(* Logix 5000 project; controller _GigaDiscovery vendor 1 type 14 code 244 rev 35.11; software revision 35.03; part 17 of 23 *)
(* tags used below, declared in another part *)
   Os : DINT;
   All_Rack_Left_Sensor_FP_OFF : BOOL;
   All_Rack_Left_Sensor_O1_OFF : BOOL;
   All_Rack_Right_Sensor_FP_OFF : BOOL;
   All_Rack_Right_Sensor_O1_OFF : BOOL;
   All_Rack_Sensor_OFF : BOOL;
   Mem_All_Rack_Sensor_OFF : BOOL;
   OS_Start_Stop_Cycle_Started : BOOL;
   Reset_Pulse : BOOL;
   RESTRAINTS_Closed : BOOL;   // All RESTRAINTS Closed
   Restraints_Cycle : Sequencer;
   RESTRAINTS_Rack : LapBar_Racks[41];
   RESTRAINTS_Rack_Sector_ON : BOOL;
   RESTRAINTS_Sector : LapBars_Sector[9];
   Start_Autom_Cycle : Sequencer;
   Start_Stop_Cycle : Sequencer;
(* S_Input, continued *)

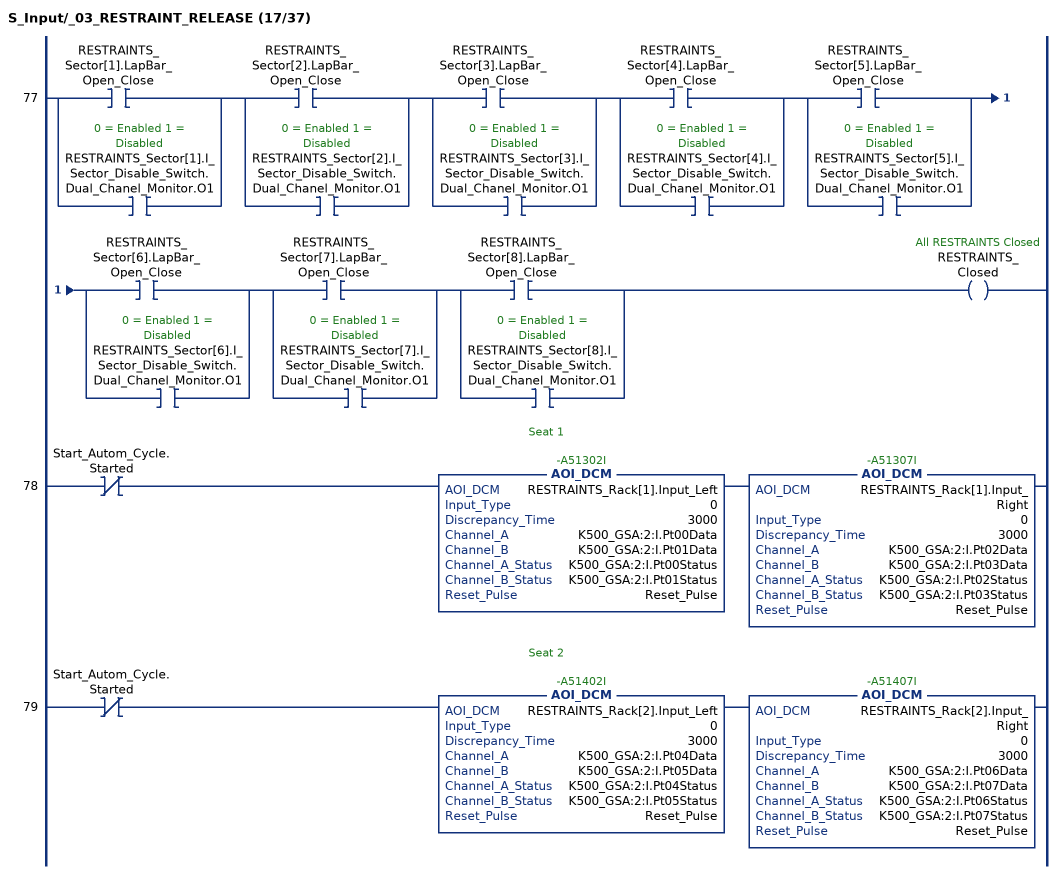
   [picture p324: S_Input/_03_RESTRAINT_RELEASE rungs 77-79]
   77: [XIC(RESTRAINTS_Sector[1].LapBar_Open_Close) ,XIC(RESTRAINTS_Sector[1].I_Sector_Disable_Switch.Dual_Chanel_Monitor.O1) ][XIC(RESTRAINTS_Sector[2].LapBar_Open_Close) ,XIC(RESTRAINTS_Sector[2].I_Sector_Disable_Switch.Dual_Chanel_Monitor.O1) ][XIC(RESTRAINTS_Sector[3].LapBar_Open_Close) ,XIC(RESTRAINTS_Sector[3].I_Sector_Disable_Switch.Dual_Chanel_Monitor.O1) ][XIC(RESTRAINTS_Sector[4].LapBar_Open_Close) ,XIC(RESTRAINTS_Sector[4].I_Sector_Disable_Switch.Dual_Chanel_Monitor.O1) ][XIC(RESTRAINTS_Sector[5].LapBar_Open_Close) ,XIC(RESTRAINTS_Sector[5].I_Sector_Disable_Switch.Dual_Chanel_Monitor.O1) ][XIC(RESTRAINTS_Sector[6].LapBar_Open_Close) ,XIC(RESTRAINTS_Sector[6].I_Sector_Disable_Switch.Dual_Chanel_Monitor.O1) ][XIC(RESTRAINTS_Sector[7].LapBar_Open_Close) ,XIC(RESTRAINTS_Sector[7].I_Sector_Disable_Switch.Dual_Chanel_Monitor.O1) ][XIC(RESTRAINTS_Sector[8].LapBar_Open_Close) ,XIC(RESTRAINTS_Sector[8].I_Sector_Disable_Switch.Dual_Chanel_Monitor.O1) ]OTE(RESTRAINTS_Closed);
   // Seat 1
   78: XIO(Start_Autom_Cycle.Started)AOI_DCM(RESTRAINTS_Rack[1].Input_Left,0,3000,K500_GSA:2:I.Pt00Data,K500_GSA:2:I.Pt01Data,K500_GSA:2:I.Pt00Status,K500_GSA:2:I.Pt01Status,Reset_Pulse)AOI_DCM(RESTRAINTS_Rack[1].Input_Right,0,3000,K500_GSA:2:I.Pt02Data,K500_GSA:2:I.Pt03Data,K500_GSA:2:I.Pt02Status,K500_GSA:2:I.Pt03Status,Reset_Pulse);
   // Seat 2
   79: XIO(Start_Autom_Cycle.Started)AOI_DCM(RESTRAINTS_Rack[2].Input_Left,0,3000,K500_GSA:2:I.Pt04Data,K500_GSA:2:I.Pt05Data,K500_GSA:2:I.Pt04Status,K500_GSA:2:I.Pt05Status,Reset_Pulse)AOI_DCM(RESTRAINTS_Rack[2].Input_Right,0,3000,K500_GSA:2:I.Pt06Data,K500_GSA:2:I.Pt07Data,K500_GSA:2:I.Pt06Status,K500_GSA:2:I.Pt07Status,Reset_Pulse);
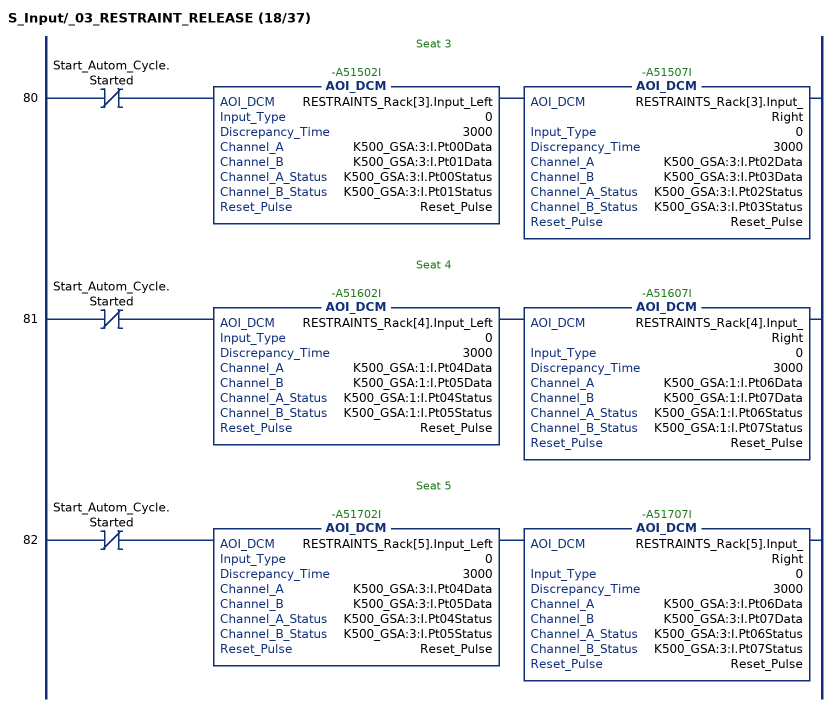
   // Seat 3
   80: XIO(Start_Autom_Cycle.Started)AOI_DCM(RESTRAINTS_Rack[3].Input_Left,0,3000,K500_GSA:3:I.Pt00Data,K500_GSA:3:I.Pt01Data,K500_GSA:3:I.Pt00Status,K500_GSA:3:I.Pt01Status,Reset_Pulse)AOI_DCM(RESTRAINTS_Rack[3].Input_Right,0,3000,K500_GSA:3:I.Pt02Data,K500_GSA:3:I.Pt03Data,K500_GSA:3:I.Pt02Status,K500_GSA:3:I.Pt03Status,Reset_Pulse);
   // Seat 4
   81: XIO(Start_Autom_Cycle.Started)AOI_DCM(RESTRAINTS_Rack[4].Input_Left,0,3000,K500_GSA:1:I.Pt04Data,K500_GSA:1:I.Pt05Data,K500_GSA:1:I.Pt04Status,K500_GSA:1:I.Pt05Status,Reset_Pulse)AOI_DCM(RESTRAINTS_Rack[4].Input_Right,0,3000,K500_GSA:1:I.Pt06Data,K500_GSA:1:I.Pt07Data,K500_GSA:1:I.Pt06Status,K500_GSA:1:I.Pt07Status,Reset_Pulse);
   // Seat 5
   82: XIO(Start_Autom_Cycle.Started)AOI_DCM(RESTRAINTS_Rack[5].Input_Left,0,3000,K500_GSA:3:I.Pt04Data,K500_GSA:3:I.Pt05Data,K500_GSA:3:I.Pt04Status,K500_GSA:3:I.Pt05Status,Reset_Pulse)AOI_DCM(RESTRAINTS_Rack[5].Input_Right,0,3000,K500_GSA:3:I.Pt06Data,K500_GSA:3:I.Pt07Data,K500_GSA:3:I.Pt06Status,K500_GSA:3:I.Pt07Status,Reset_Pulse);
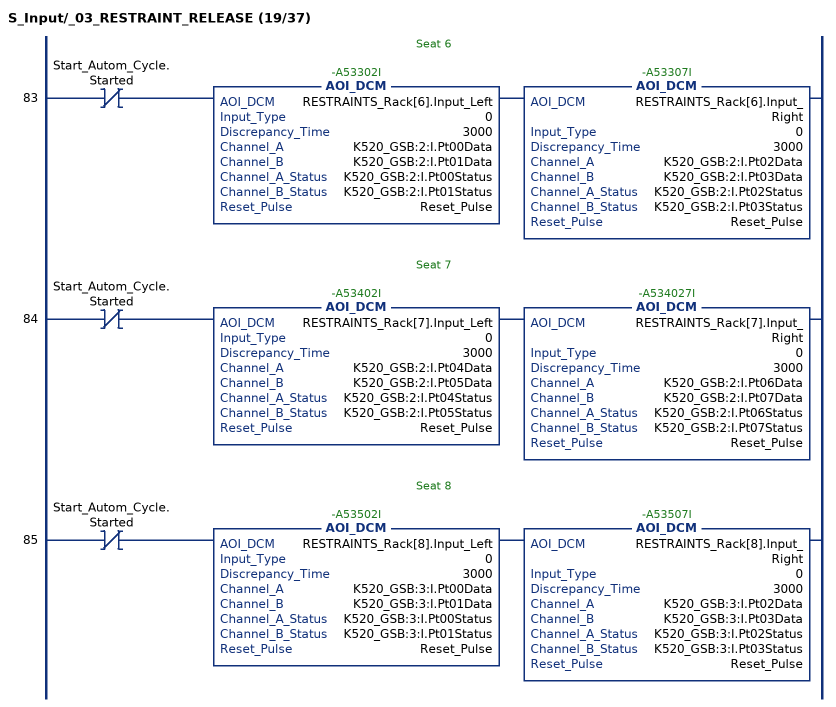
   // Seat 6
   83: XIO(Start_Autom_Cycle.Started)AOI_DCM(RESTRAINTS_Rack[6].Input_Left,0,3000,K520_GSB:2:I.Pt00Data,K520_GSB:2:I.Pt01Data,K520_GSB:2:I.Pt00Status,K520_GSB:2:I.Pt01Status,Reset_Pulse)AOI_DCM(RESTRAINTS_Rack[6].Input_Right,0,3000,K520_GSB:2:I.Pt02Data,K520_GSB:2:I.Pt03Data,K520_GSB:2:I.Pt02Status,K520_GSB:2:I.Pt03Status,Reset_Pulse);
   // Seat 7
   84: XIO(Start_Autom_Cycle.Started)AOI_DCM(RESTRAINTS_Rack[7].Input_Left,0,3000,K520_GSB:2:I.Pt04Data,K520_GSB:2:I.Pt05Data,K520_GSB:2:I.Pt04Status,K520_GSB:2:I.Pt05Status,Reset_Pulse)AOI_DCM(RESTRAINTS_Rack[7].Input_Right,0,3000,K520_GSB:2:I.Pt06Data,K520_GSB:2:I.Pt07Data,K520_GSB:2:I.Pt06Status,K520_GSB:2:I.Pt07Status,Reset_Pulse);
   // Seat 8
   85: XIO(Start_Autom_Cycle.Started)AOI_DCM(RESTRAINTS_Rack[8].Input_Left,0,3000,K520_GSB:3:I.Pt00Data,K520_GSB:3:I.Pt01Data,K520_GSB:3:I.Pt00Status,K520_GSB:3:I.Pt01Status,Reset_Pulse)AOI_DCM(RESTRAINTS_Rack[8].Input_Right,0,3000,K520_GSB:3:I.Pt02Data,K520_GSB:3:I.Pt03Data,K520_GSB:3:I.Pt02Status,K520_GSB:3:I.Pt03Status,Reset_Pulse);
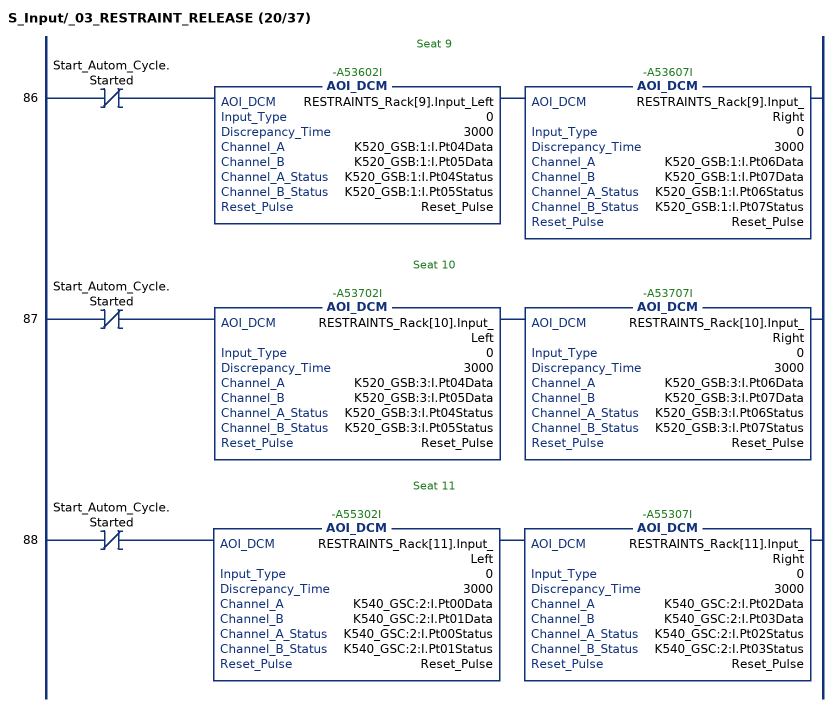
   // Seat 9
   86: XIO(Start_Autom_Cycle.Started)AOI_DCM(RESTRAINTS_Rack[9].Input_Left,0,3000,K520_GSB:1:I.Pt04Data,K520_GSB:1:I.Pt05Data,K520_GSB:1:I.Pt04Status,K520_GSB:1:I.Pt05Status,Reset_Pulse)AOI_DCM(RESTRAINTS_Rack[9].Input_Right,0,3000,K520_GSB:1:I.Pt06Data,K520_GSB:1:I.Pt07Data,K520_GSB:1:I.Pt06Status,K520_GSB:1:I.Pt07Status,Reset_Pulse);
   // Seat 10
   87: XIO(Start_Autom_Cycle.Started)AOI_DCM(RESTRAINTS_Rack[10].Input_Left,0,3000,K520_GSB:3:I.Pt04Data,K520_GSB:3:I.Pt05Data,K520_GSB:3:I.Pt04Status,K520_GSB:3:I.Pt05Status,Reset_Pulse)AOI_DCM(RESTRAINTS_Rack[10].Input_Right,0,3000,K520_GSB:3:I.Pt06Data,K520_GSB:3:I.Pt07Data,K520_GSB:3:I.Pt06Status,K520_GSB:3:I.Pt07Status,Reset_Pulse);
   // Seat 11
   88: XIO(Start_Autom_Cycle.Started)AOI_DCM(RESTRAINTS_Rack[11].Input_Left,0,3000,K540_GSC:2:I.Pt00Data,K540_GSC:2:I.Pt01Data,K540_GSC:2:I.Pt00Status,K540_GSC:2:I.Pt01Status,Reset_Pulse)AOI_DCM(RESTRAINTS_Rack[11].Input_Right,0,3000,K540_GSC:2:I.Pt02Data,K540_GSC:2:I.Pt03Data,K540_GSC:2:I.Pt02Status,K540_GSC:2:I.Pt03Status,Reset_Pulse);
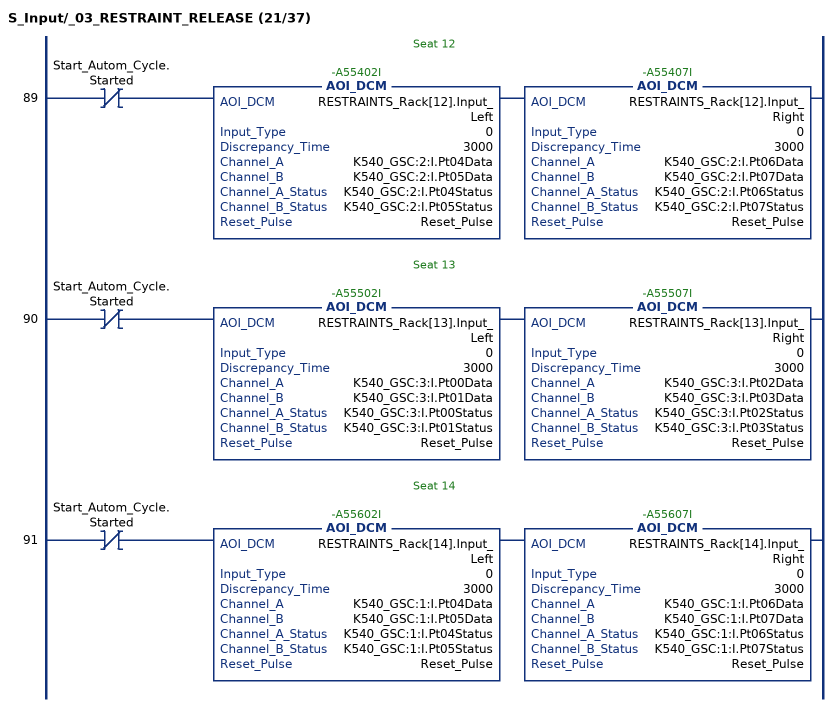
   // Seat 12
   89: XIO(Start_Autom_Cycle.Started)AOI_DCM(RESTRAINTS_Rack[12].Input_Left,0,3000,K540_GSC:2:I.Pt04Data,K540_GSC:2:I.Pt05Data,K540_GSC:2:I.Pt04Status,K540_GSC:2:I.Pt05Status,Reset_Pulse)AOI_DCM(RESTRAINTS_Rack[12].Input_Right,0,3000,K540_GSC:2:I.Pt06Data,K540_GSC:2:I.Pt07Data,K540_GSC:2:I.Pt06Status,K540_GSC:2:I.Pt07Status,Reset_Pulse);
   // Seat 13
   90: XIO(Start_Autom_Cycle.Started)AOI_DCM(RESTRAINTS_Rack[13].Input_Left,0,3000,K540_GSC:3:I.Pt00Data,K540_GSC:3:I.Pt01Data,K540_GSC:3:I.Pt00Status,K540_GSC:3:I.Pt01Status,Reset_Pulse)AOI_DCM(RESTRAINTS_Rack[13].Input_Right,0,3000,K540_GSC:3:I.Pt02Data,K540_GSC:3:I.Pt03Data,K540_GSC:3:I.Pt02Status,K540_GSC:3:I.Pt03Status,Reset_Pulse);
   // Seat 14
   91: XIO(Start_Autom_Cycle.Started)AOI_DCM(RESTRAINTS_Rack[14].Input_Left,0,3000,K540_GSC:1:I.Pt04Data,K540_GSC:1:I.Pt05Data,K540_GSC:1:I.Pt04Status,K540_GSC:1:I.Pt05Status,Reset_Pulse)AOI_DCM(RESTRAINTS_Rack[14].Input_Right,0,3000,K540_GSC:1:I.Pt06Data,K540_GSC:1:I.Pt07Data,K540_GSC:1:I.Pt06Status,K540_GSC:1:I.Pt07Status,Reset_Pulse);
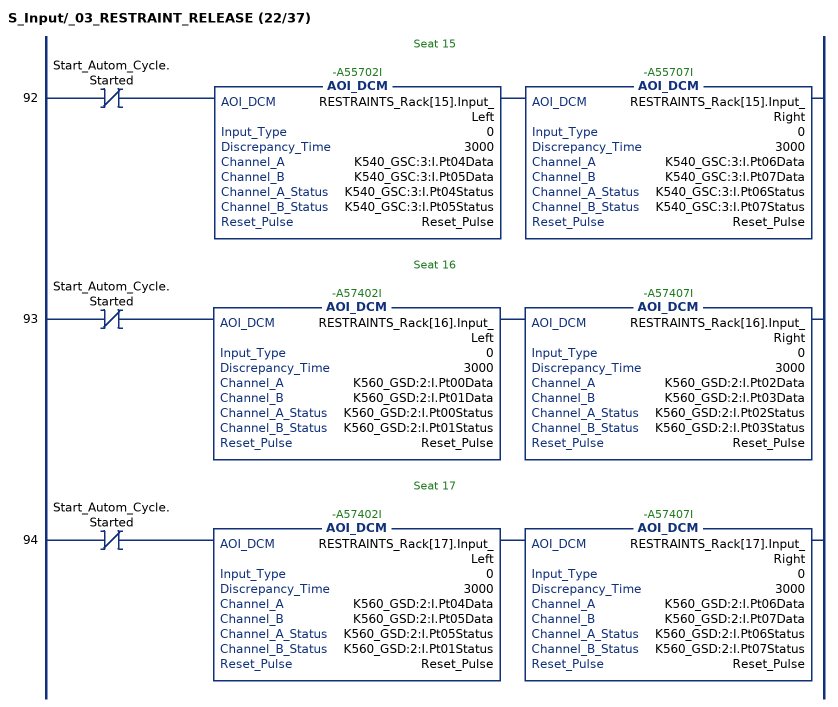
   // Seat 15
   92: XIO(Start_Autom_Cycle.Started)AOI_DCM(RESTRAINTS_Rack[15].Input_Left,0,3000,K540_GSC:3:I.Pt04Data,K540_GSC:3:I.Pt05Data,K540_GSC:3:I.Pt04Status,K540_GSC:3:I.Pt05Status,Reset_Pulse)AOI_DCM(RESTRAINTS_Rack[15].Input_Right,0,3000,K540_GSC:3:I.Pt06Data,K540_GSC:3:I.Pt07Data,K540_GSC:3:I.Pt06Status,K540_GSC:3:I.Pt07Status,Reset_Pulse);
   // Seat 16
   93: XIO(Start_Autom_Cycle.Started)AOI_DCM(RESTRAINTS_Rack[16].Input_Left,0,3000,K560_GSD:2:I.Pt00Data,K560_GSD:2:I.Pt01Data,K560_GSD:2:I.Pt00Status,K560_GSD:2:I.Pt01Status,Reset_Pulse)AOI_DCM(RESTRAINTS_Rack[16].Input_Right,0,3000,K560_GSD:2:I.Pt02Data,K560_GSD:2:I.Pt03Data,K560_GSD:2:I.Pt02Status,K560_GSD:2:I.Pt03Status,Reset_Pulse);
   // Seat 17
   94: XIO(Start_Autom_Cycle.Started)AOI_DCM(RESTRAINTS_Rack[17].Input_Left,0,3000,K560_GSD:2:I.Pt04Data,K560_GSD:2:I.Pt05Data,K560_GSD:2:I.Pt05Status,K560_GSD:2:I.Pt01Status,Reset_Pulse)AOI_DCM(RESTRAINTS_Rack[17].Input_Right,0,3000,K560_GSD:2:I.Pt06Data,K560_GSD:2:I.Pt07Data,K560_GSD:2:I.Pt06Status,K560_GSD:2:I.Pt07Status,Reset_Pulse);
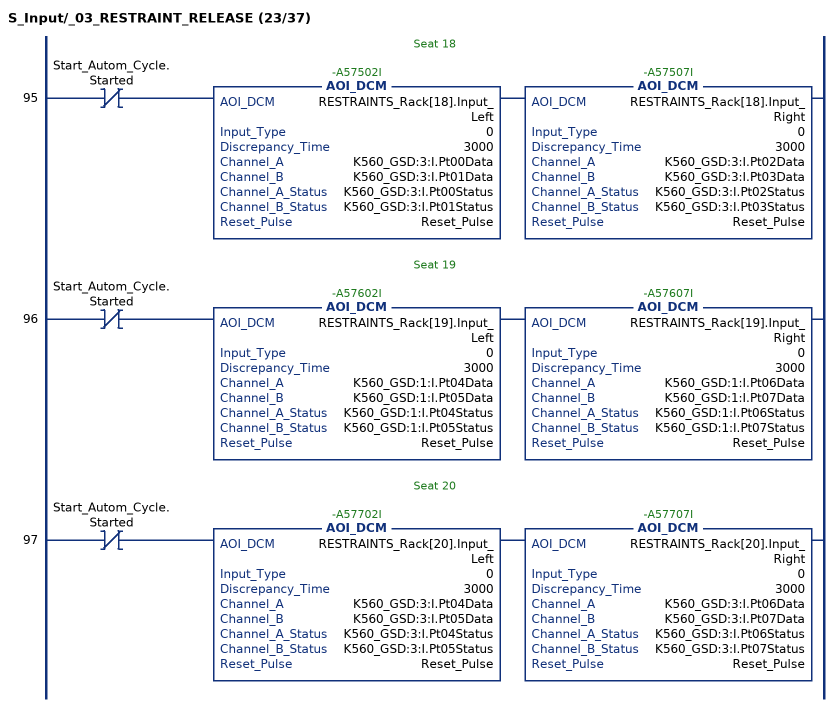
   // Seat 18
   95: XIO(Start_Autom_Cycle.Started)AOI_DCM(RESTRAINTS_Rack[18].Input_Left,0,3000,K560_GSD:3:I.Pt00Data,K560_GSD:3:I.Pt01Data,K560_GSD:3:I.Pt00Status,K560_GSD:3:I.Pt01Status,Reset_Pulse)AOI_DCM(RESTRAINTS_Rack[18].Input_Right,0,3000,K560_GSD:3:I.Pt02Data,K560_GSD:3:I.Pt03Data,K560_GSD:3:I.Pt02Status,K560_GSD:3:I.Pt03Status,Reset_Pulse);
   // Seat 19
   96: XIO(Start_Autom_Cycle.Started)AOI_DCM(RESTRAINTS_Rack[19].Input_Left,0,3000,K560_GSD:1:I.Pt04Data,K560_GSD:1:I.Pt05Data,K560_GSD:1:I.Pt04Status,K560_GSD:1:I.Pt05Status,Reset_Pulse)AOI_DCM(RESTRAINTS_Rack[19].Input_Right,0,3000,K560_GSD:1:I.Pt06Data,K560_GSD:1:I.Pt07Data,K560_GSD:1:I.Pt06Status,K560_GSD:1:I.Pt07Status,Reset_Pulse);
   // Seat 20
   97: XIO(Start_Autom_Cycle.Started)AOI_DCM(RESTRAINTS_Rack[20].Input_Left,0,3000,K560_GSD:3:I.Pt04Data,K560_GSD:3:I.Pt05Data,K560_GSD:3:I.Pt04Status,K560_GSD:3:I.Pt05Status,Reset_Pulse)AOI_DCM(RESTRAINTS_Rack[20].Input_Right,0,3000,K560_GSD:3:I.Pt06Data,K560_GSD:3:I.Pt07Data,K560_GSD:3:I.Pt06Status,K560_GSD:3:I.Pt07Status,Reset_Pulse);
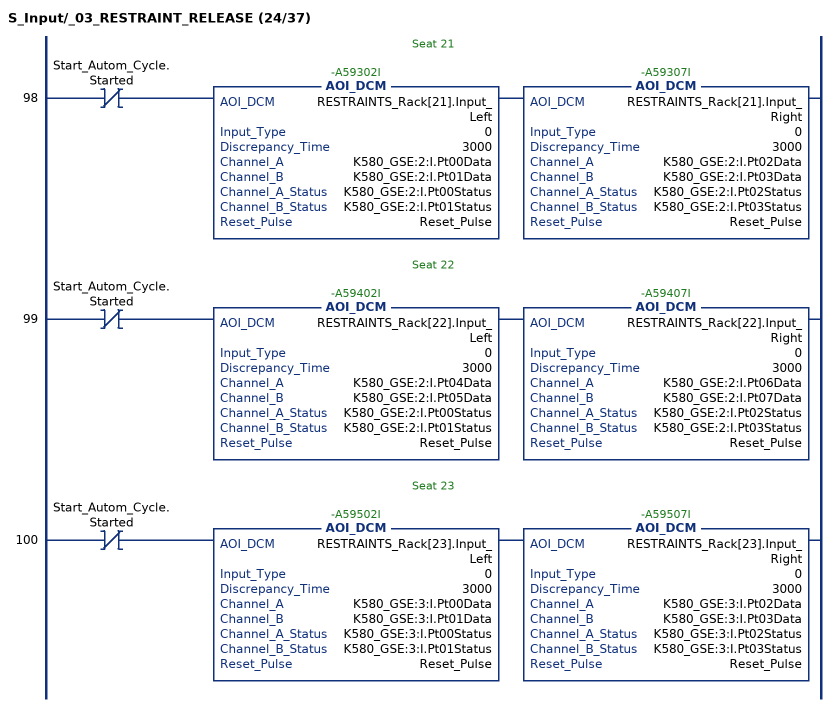
   // Seat 21
   98: XIO(Start_Autom_Cycle.Started)AOI_DCM(RESTRAINTS_Rack[21].Input_Left,0,3000,K580_GSE:2:I.Pt00Data,K580_GSE:2:I.Pt01Data,K580_GSE:2:I.Pt00Status,K580_GSE:2:I.Pt01Status,Reset_Pulse)AOI_DCM(RESTRAINTS_Rack[21].Input_Right,0,3000,K580_GSE:2:I.Pt02Data,K580_GSE:2:I.Pt03Data,K580_GSE:2:I.Pt02Status,K580_GSE:2:I.Pt03Status,Reset_Pulse);
   // Seat 22
   99: XIO(Start_Autom_Cycle.Started)AOI_DCM(RESTRAINTS_Rack[22].Input_Left,0,3000,K580_GSE:2:I.Pt04Data,K580_GSE:2:I.Pt05Data,K580_GSE:2:I.Pt00Status,K580_GSE:2:I.Pt01Status,Reset_Pulse)AOI_DCM(RESTRAINTS_Rack[22].Input_Right,0,3000,K580_GSE:2:I.Pt06Data,K580_GSE:2:I.Pt07Data,K580_GSE:2:I.Pt02Status,K580_GSE:2:I.Pt03Status,Reset_Pulse);
   // Seat 23
   100: XIO(Start_Autom_Cycle.Started)AOI_DCM(RESTRAINTS_Rack[23].Input_Left,0,3000,K580_GSE:3:I.Pt00Data,K580_GSE:3:I.Pt01Data,K580_GSE:3:I.Pt00Status,K580_GSE:3:I.Pt01Status,Reset_Pulse)AOI_DCM(RESTRAINTS_Rack[23].Input_Right,0,3000,K580_GSE:3:I.Pt02Data,K580_GSE:3:I.Pt03Data,K580_GSE:3:I.Pt02Status,K580_GSE:3:I.Pt03Status,Reset_Pulse);
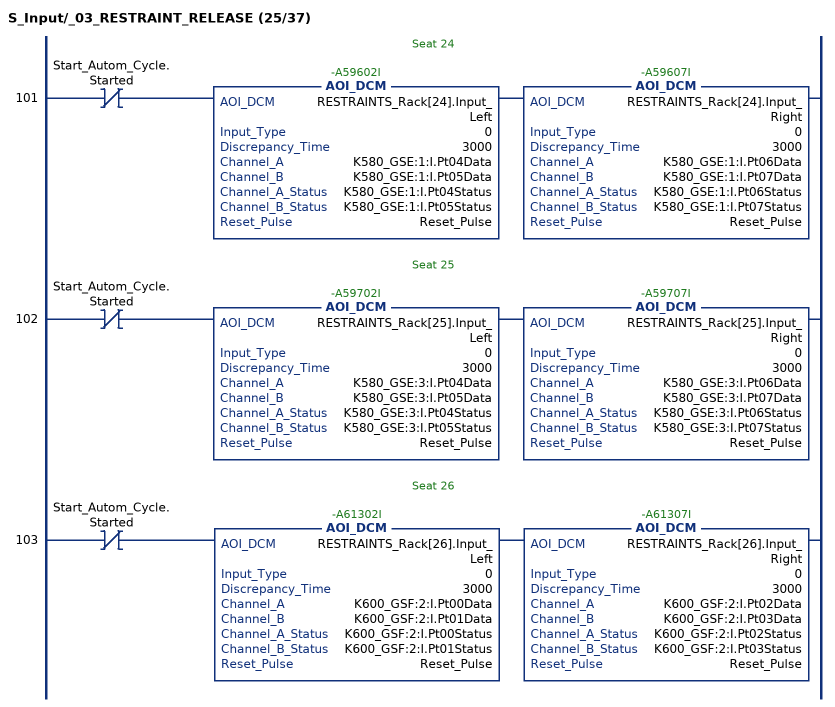
   // Seat 24
   101: XIO(Start_Autom_Cycle.Started)AOI_DCM(RESTRAINTS_Rack[24].Input_Left,0,3000,K580_GSE:1:I.Pt04Data,K580_GSE:1:I.Pt05Data,K580_GSE:1:I.Pt04Status,K580_GSE:1:I.Pt05Status,Reset_Pulse)AOI_DCM(RESTRAINTS_Rack[24].Input_Right,0,3000,K580_GSE:1:I.Pt06Data,K580_GSE:1:I.Pt07Data,K580_GSE:1:I.Pt06Status,K580_GSE:1:I.Pt07Status,Reset_Pulse);
   // Seat 25
   102: XIO(Start_Autom_Cycle.Started)AOI_DCM(RESTRAINTS_Rack[25].Input_Left,0,3000,K580_GSE:3:I.Pt04Data,K580_GSE:3:I.Pt05Data,K580_GSE:3:I.Pt04Status,K580_GSE:3:I.Pt05Status,Reset_Pulse)AOI_DCM(RESTRAINTS_Rack[25].Input_Right,0,3000,K580_GSE:3:I.Pt06Data,K580_GSE:3:I.Pt07Data,K580_GSE:3:I.Pt06Status,K580_GSE:3:I.Pt07Status,Reset_Pulse);
   // Seat 26
   103: XIO(Start_Autom_Cycle.Started)AOI_DCM(RESTRAINTS_Rack[26].Input_Left,0,3000,K600_GSF:2:I.Pt00Data,K600_GSF:2:I.Pt01Data,K600_GSF:2:I.Pt00Status,K600_GSF:2:I.Pt01Status,Reset_Pulse)AOI_DCM(RESTRAINTS_Rack[26].Input_Right,0,3000,K600_GSF:2:I.Pt02Data,K600_GSF:2:I.Pt03Data,K600_GSF:2:I.Pt02Status,K600_GSF:2:I.Pt03Status,Reset_Pulse);
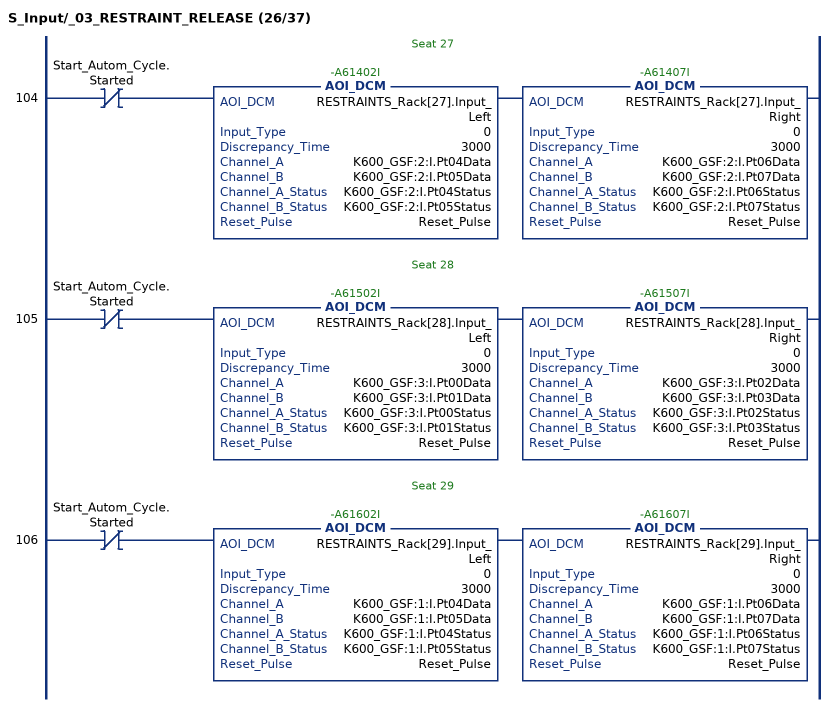
   // Seat 27
   104: XIO(Start_Autom_Cycle.Started)AOI_DCM(RESTRAINTS_Rack[27].Input_Left,0,3000,K600_GSF:2:I.Pt04Data,K600_GSF:2:I.Pt05Data,K600_GSF:2:I.Pt04Status,K600_GSF:2:I.Pt05Status,Reset_Pulse)AOI_DCM(RESTRAINTS_Rack[27].Input_Right,0,3000,K600_GSF:2:I.Pt06Data,K600_GSF:2:I.Pt07Data,K600_GSF:2:I.Pt06Status,K600_GSF:2:I.Pt07Status,Reset_Pulse);
   // Seat 28
   105: XIO(Start_Autom_Cycle.Started)AOI_DCM(RESTRAINTS_Rack[28].Input_Left,0,3000,K600_GSF:3:I.Pt00Data,K600_GSF:3:I.Pt01Data,K600_GSF:3:I.Pt00Status,K600_GSF:3:I.Pt01Status,Reset_Pulse)AOI_DCM(RESTRAINTS_Rack[28].Input_Right,0,3000,K600_GSF:3:I.Pt02Data,K600_GSF:3:I.Pt03Data,K600_GSF:3:I.Pt02Status,K600_GSF:3:I.Pt03Status,Reset_Pulse);
   // Seat 29
   106: XIO(Start_Autom_Cycle.Started)AOI_DCM(RESTRAINTS_Rack[29].Input_Left,0,3000,K600_GSF:1:I.Pt04Data,K600_GSF:1:I.Pt05Data,K600_GSF:1:I.Pt04Status,K600_GSF:1:I.Pt05Status,Reset_Pulse)AOI_DCM(RESTRAINTS_Rack[29].Input_Right,0,3000,K600_GSF:1:I.Pt06Data,K600_GSF:1:I.Pt07Data,K600_GSF:1:I.Pt06Status,K600_GSF:1:I.Pt07Status,Reset_Pulse);
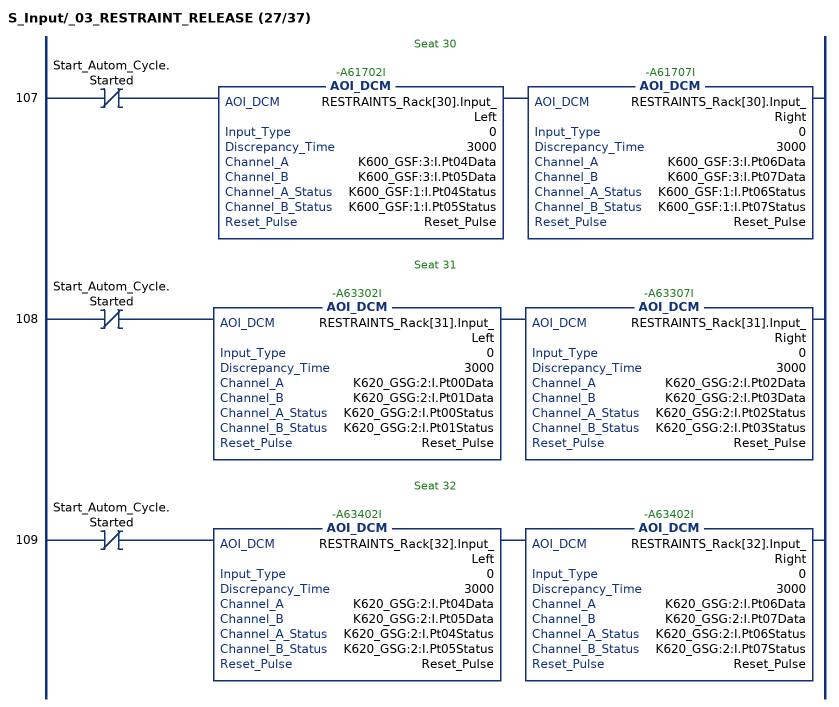
   // Seat 30
   107: XIO(Start_Autom_Cycle.Started)AOI_DCM(RESTRAINTS_Rack[30].Input_Left,0,3000,K600_GSF:3:I.Pt04Data,K600_GSF:3:I.Pt05Data,K600_GSF:1:I.Pt04Status,K600_GSF:1:I.Pt05Status,Reset_Pulse)AOI_DCM(RESTRAINTS_Rack[30].Input_Right,0,3000,K600_GSF:3:I.Pt06Data,K600_GSF:3:I.Pt07Data,K600_GSF:1:I.Pt06Status,K600_GSF:1:I.Pt07Status,Reset_Pulse);
   // Seat 31
   108: XIO(Start_Autom_Cycle.Started)AOI_DCM(RESTRAINTS_Rack[31].Input_Left,0,3000,K620_GSG:2:I.Pt00Data,K620_GSG:2:I.Pt01Data,K620_GSG:2:I.Pt00Status,K620_GSG:2:I.Pt01Status,Reset_Pulse)AOI_DCM(RESTRAINTS_Rack[31].Input_Right,0,3000,K620_GSG:2:I.Pt02Data,K620_GSG:2:I.Pt03Data,K620_GSG:2:I.Pt02Status,K620_GSG:2:I.Pt03Status,Reset_Pulse);
   // Seat 32
   109: XIO(Start_Autom_Cycle.Started)AOI_DCM(RESTRAINTS_Rack[32].Input_Left,0,3000,K620_GSG:2:I.Pt04Data,K620_GSG:2:I.Pt05Data,K620_GSG:2:I.Pt04Status,K620_GSG:2:I.Pt05Status,Reset_Pulse)AOI_DCM(RESTRAINTS_Rack[32].Input_Right,0,3000,K620_GSG:2:I.Pt06Data,K620_GSG:2:I.Pt07Data,K620_GSG:2:I.Pt06Status,K620_GSG:2:I.Pt07Status,Reset_Pulse);
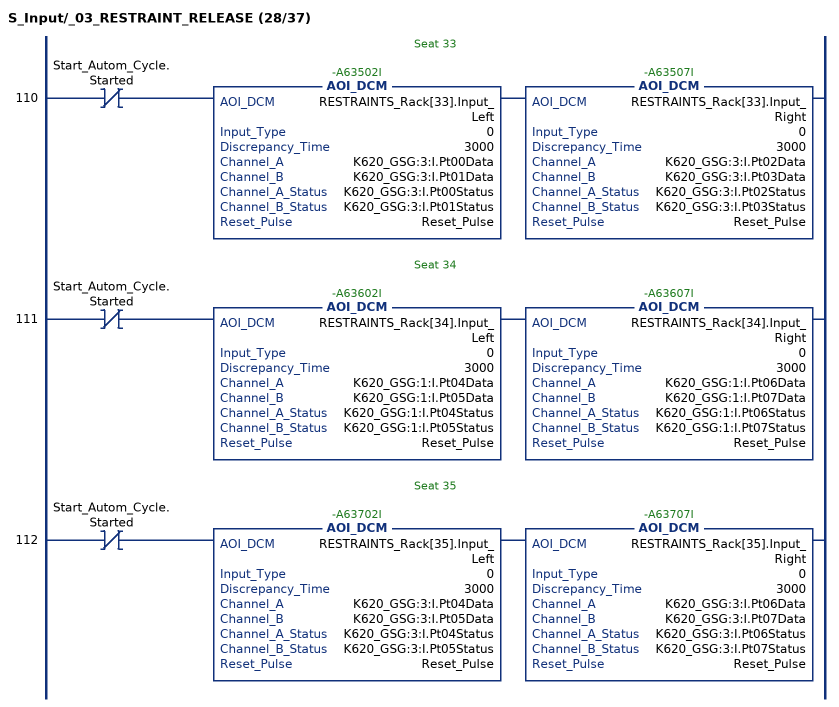
   // Seat 33
   110: XIO(Start_Autom_Cycle.Started)AOI_DCM(RESTRAINTS_Rack[33].Input_Left,0,3000,K620_GSG:3:I.Pt00Data,K620_GSG:3:I.Pt01Data,K620_GSG:3:I.Pt00Status,K620_GSG:3:I.Pt01Status,Reset_Pulse)AOI_DCM(RESTRAINTS_Rack[33].Input_Right,0,3000,K620_GSG:3:I.Pt02Data,K620_GSG:3:I.Pt03Data,K620_GSG:3:I.Pt02Status,K620_GSG:3:I.Pt03Status,Reset_Pulse);
   // Seat 34
   111: XIO(Start_Autom_Cycle.Started)AOI_DCM(RESTRAINTS_Rack[34].Input_Left,0,3000,K620_GSG:1:I.Pt04Data,K620_GSG:1:I.Pt05Data,K620_GSG:1:I.Pt04Status,K620_GSG:1:I.Pt05Status,Reset_Pulse)AOI_DCM(RESTRAINTS_Rack[34].Input_Right,0,3000,K620_GSG:1:I.Pt06Data,K620_GSG:1:I.Pt07Data,K620_GSG:1:I.Pt06Status,K620_GSG:1:I.Pt07Status,Reset_Pulse);
   // Seat 35
   112: XIO(Start_Autom_Cycle.Started)AOI_DCM(RESTRAINTS_Rack[35].Input_Left,0,3000,K620_GSG:3:I.Pt04Data,K620_GSG:3:I.Pt05Data,K620_GSG:3:I.Pt04Status,K620_GSG:3:I.Pt05Status,Reset_Pulse)AOI_DCM(RESTRAINTS_Rack[35].Input_Right,0,3000,K620_GSG:3:I.Pt06Data,K620_GSG:3:I.Pt07Data,K620_GSG:3:I.Pt06Status,K620_GSG:3:I.Pt07Status,Reset_Pulse);